REGION Network 23: Buzzer
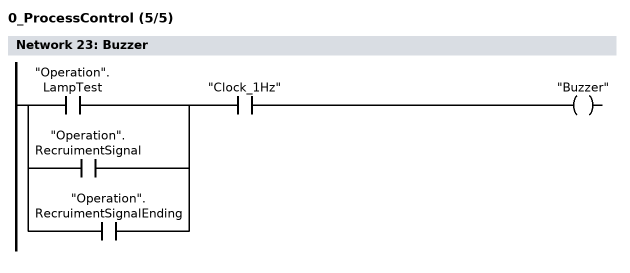
   RUNG wire#powerrail
      Contact( "Operation".LampTest )
      wire#w1
      Contact( "Clock_1Hz" )
      Coil( "Buzzer" )
   END_RUNG
   RUNG wire#powerrail
      Contact( "Operation".RecruimentSignal )
   END_RUNG wire#w1
   RUNG wire#powerrail
      Contact( "Operation".RecruimentSignalEnding )
   END_RUNG wire#w1
   // the same network as SCL:
   "Buzzer" := ("Operation".LampTest OR "Operation".RecruimentSignal OR "Operation".RecruimentSignalEnding) AND "Clock_1Hz";
END_REGION
END_FUNCTION_BLOCK

// folder: 5_Library

FUNCTION_BLOCK "DigAlarm"   // FB2000, SCL
TITLE = Digital Alarm
{ S7_Optimized_Access := 'TRUE' }
AUTHOR : JL_Cristobal_2020
VERSION : 0.1
// Digital Alarm supervisor, trigger memory , ack + reset
   VAR_INPUT
      Pulse : Bool;
      ACK : Bool;
      Reset : Bool;
      Funtion : Bool;
      Input : Bool;
   END_VAR
   VAR_OUTPUT
      DisplayOutput : Bool;
      DisplayOutputNeg : Bool;
      InterlockOutput : Bool;
      InterlockOutputNeg : Bool;
   END_VAR
   VAR
      DisplayAlarmMem : Bool;
      ACKMem : Bool;
      InterlockalarmMem : Bool;
      InterlockMem : Bool;
   END_VAR
BEGIN
   //Alarm process

   //TRUE Mode, Positive Signal
   IF #Funtion = 1 THEN

       IF NOT #Input THEN
           #InterlockMem := false;
           #DisplayAlarmMem := true;
           #InterlockalarmMem := true;
       END_IF;

       IF #Input AND #Reset THEN
           #DisplayAlarmMem := false;
       END_IF;

       IF NOT #Input AND #ACK THEN
           #ACKMem := true;
       END_IF;

       IF #Input AND #Reset THEN
           #InterlockMem := true;
           #ACKMem := false;
           #InterlockalarmMem := false;
       END_IF;

   END_IF;

   //FALSE Mode, Negative Signal
   IF #Funtion = 0 THEN

       IF #Input THEN
           #DisplayAlarmMem := true;
           #InterlockalarmMem := true;
           #InterlockMem := false;
       END_IF;

       IF NOT #Input AND #Reset THEN
           #DisplayAlarmMem := false;
       END_IF;

       IF #Input AND #ACK THEN
           #ACKMem := true;
       END_IF;

       IF NOT #Input AND #Reset THEN
           #ACKMem := false;
           #InterlockalarmMem := false;
           #InterlockMem := true;
       END_IF;

   END_IF;


   #DisplayOutput := #DisplayAlarmMem AND ((#Pulse AND NOT #ACKMem) OR #ACKMem);
   #DisplayOutputNeg := NOT (#DisplayAlarmMem AND ((#Pulse AND NOT #ACKMem) OR #ACKMem));
   #InterlockOutput := #InterlockMem;
   #InterlockOutputNeg := NOT #InterlockMem;
END_FUNCTION_BLOCK

FUNCTION_BLOCK "DigAlarmInterlock"   // FB2001, SCL
TITLE = Digital Alarm With Interlock
{ S7_Optimized_Access := 'TRUE' }
AUTHOR : JL_Cristobal_2020
FAMILY : Alarms
VERSION : 0.1
// Digital Alarm supervisor with interlock signal, trigger memory , ack + reset
   VAR_INPUT
      Pulse : Bool;
      ACK : Bool;
      Reset : Bool;
      Function : Int;
      AlarmInput : Bool;
      SupervisorInput : Bool;
      StartInput : Bool;
      Delay : Time;
   END_VAR
   VAR_OUTPUT
      DisplayOutput : Bool;
      DisplayOutputNeg : Bool;
      InterlockOutput : Bool;
      InterlockOutputNeg : Bool;
      SupervisorOutput : Bool;
      TimeElapsed : Time;
   END_VAR
   VAR RETAIN
      DisplayAlarmMem : Bool;
      ACKMem : Bool;
      InterlockalarmMem : Bool;
      InterlockMem : Bool;
   END_VAR
   VAR
      EndSPVMem : Bool;
   END_VAR
   VAR RETAIN
      SPVMem : Bool;
   END_VAR
BEGIN
   (*GESTION DE LA ALARMA*)

   //TRUE MODE, ACTIVE OK
   IF #Function = 1 OR #Function=3 THEN

       IF NOT #AlarmInput THEN
           #InterlockMem := false;
           #DisplayAlarmMem := true;
           #InterlockalarmMem := true;
       END_IF;

       IF #AlarmInput AND #Reset THEN
           #DisplayAlarmMem := false;
       END_IF;

       IF NOT #AlarmInput AND #ACK THEN
           #ACKMem := true;
       END_IF;

       IF #AlarmInput AND #Reset THEN
           #InterlockMem := true;
           #ACKMem := false;
           #InterlockalarmMem := false;
       END_IF;

   END_IF;

   //FALSE MODE, PASIVE OK
   IF #Function = 0 OR #Function=2 THEN

       IF #AlarmInput THEN
           #DisplayAlarmMem := true;
           #InterlockalarmMem := true;
           #InterlockMem := false;
       END_IF;

       IF NOT #AlarmInput AND #Reset THEN
           #DisplayAlarmMem := false;
       END_IF;

       IF #AlarmInput AND #ACK THEN
           #ACKMem := true;
       END_IF;

       IF NOT #AlarmInput AND #Reset THEN
           #ACKMem := false;
           #InterlockalarmMem := false;
           #InterlockMem := true;
       END_IF;
   END_IF;

   //SUPERVISION CONTROL
   IF #Function = 0 OR #Function = 1 THEN
       IF #StartInput THEN
           "IEC_Timer_0_DB_SPV".TON(IN := #StartInput,
                                    PT := #Delay,
                                    Q => #EndSPVMem,
                                    ET => #TimeElapsed);
           IF #EndSPVMem AND NOT #SupervisorInput THEN
               #SPVMem := 1;
           END_IF;
       ELSE
           #SPVMem := 0;
       END_IF;
   END_IF;


   #DisplayOutput := #DisplayAlarmMem AND ((#Pulse AND NOT #ACKMem) OR #ACKMem);
   #DisplayOutputNeg := NOT (#DisplayAlarmMem AND ((#Pulse AND NOT #ACKMem) OR #ACKMem));
   #InterlockOutput := #InterlockMem;
   #InterlockOutputNeg := NOT #InterlockMem;
END_FUNCTION_BLOCK

FUNCTION_BLOCK "DirectAnalog"   // FB2002, SCL
TITLE = Analog Alarm INT
{ S7_Optimized_Access := 'FALSE' }
AUTHOR : JL_Cristobal_2020
VERSION : 0.1
// Analog (int) Alarm supervisor, trigger memory , ack + reset. Prealarm and alarm for HI and LOW levels
   VAR_INPUT
      Pulse : Bool;
      ACK : Bool;
      Reset : Bool;
      Interlock : Bool;
      Delay : Time;
      Factor : Real;
      AnalogInput : Int;
      SetpointPreAlarmHI : Real;
      SetpointAlarmHI : Real;
      SetpointPreAlarmLOW : Real;
      SetpointAlarmLOW : Real;
      HysteresisHI : Real;
      HysteresisLOW : Real;
   END_VAR
   VAR_OUTPUT
      DisplayPreAlarmHI : Bool;
      InterlockPreAlarmHI : Bool;
      DisplayAlarmHI : Bool;
      InterlockAlarmHI : Bool;
      DisplayPreAlarmLOW : Bool;
      InterlockPreAlarmLOW : Bool;
      DisplayAlarmLOW : Bool;
      InterlockAlarmLOW : Bool;
      CovertedOutput : Real;
      CalcHysterisHI : Real;
      CalcHysteresisLOW : Real;
      DATOS : Struct
         InterlockPreAlarmHI : Bool;
         InterlockAlarmHI : Bool;
         InterlockPreAlarmLOW : Bool;
         InterlockAlarmLOW : Bool;
         CovertedOutput : Real;
         Error : Bool;
      END_STRUCT;
   END_VAR
   VAR
      MemDisplayPreAlarmHI : Bool;
      MemInterlockPreAlarmHI : Bool;
      MemDisplayAlarmHI : Bool;
      MemInterlockAlarmHI : Bool;
      MemDisplayPreAlarmLOW : Bool;
      MemInterlockPreAlarmLOW : Bool;
      MemDisplayAlarmLOW : Bool;
      MemInterlockAlarmLOW : Bool;
   END_VAR
BEGIN
   //Unit conversion
   #CovertedOutput := #AnalogInput/#Factor;

   //Prealarm HI
   //Set PreAlarm
   IF #Interlock AND (#CovertedOutput >= #SetpointPreAlarmHI) THEN
     #InterlockPreAlarmHI := false;
     #MemDisplayPreAlarmHI := true;
   END_IF;
   //ACK
   IF (#MemDisplayPreAlarmHI OR NOT #MemInterlockPreAlarmHI) AND #ACK THEN
     #MemInterlockPreAlarmHI := true;
   END_IF;
   //Reset
   IF(#CovertedOutput < (#SetpointPreAlarmHI - #HysteresisHI)) THEN
     #InterlockPreAlarmHI := true;
     #MemDisplayPreAlarmHI := false;
     #MemInterlockPreAlarmHI := false;
   END_IF;
   //Display Output
   #DisplayPreAlarmHI := NOT #InterlockPreAlarmHI AND ((#Pulse AND NOT #MemInterlockPreAlarmHI) OR #MemInterlockPreAlarmHI);

   //Alarm HI
   //Set Alarm HI
   IF #Interlock AND (#CovertedOutput >= #SetpointAlarmHI) THEN
       #InterlockAlarmHI := false;
     #MemDisplayAlarmHI := true;
   END_IF;
   //ACK
   IF (#MemDisplayAlarmHI OR NOT #MemInterlockAlarmHI) AND #ACK THEN
     #MemInterlockAlarmHI := true;
   END_IF;
   //Reset
   IF(#CovertedOutput < (#SetpointAlarmHI - #HysteresisHI)) THEN
     #InterlockAlarmHI := true;
     #MemDisplayAlarmHI := false;
     #MemInterlockAlarmHI := false;
   END_IF;
   //Display Output
   #DisplayAlarmHI := NOT #InterlockAlarmHI AND ((#Pulse AND NOT #MemInterlockAlarmHI) OR #MemInterlockAlarmHI);
   #CalcHysterisHI := #SetpointAlarmHI - #HysteresisHI;

   //Prealarm LOW
   //Set PreAlarm LOW
   IF #Interlock AND (#CovertedOutput <= #SetpointPreAlarmLOW) THEN
     #InterlockPreAlarmLOW := false;
     #MemDisplayPreAlarmLOW := true;
   END_IF;
   //ACK
   IF (#MemDisplayPreAlarmLOW OR NOT #MemInterlockPreAlarmLOW) AND #ACK THEN
     #MemInterlockPreAlarmLOW := true;
   END_IF;
   //Reset
   IF (#CovertedOutput > (#SetpointPreAlarmLOW + #HysteresisLOW)) THEN
     #InterlockPreAlarmLOW := true;
     #MemDisplayPreAlarmLOW := false;
     #MemInterlockPreAlarmLOW := false;
   END_IF;
   //Display Output
   #DisplayPreAlarmLOW := NOT #InterlockPreAlarmLOW AND ((#Pulse AND NOT #MemInterlockPreAlarmLOW) OR #MemInterlockPreAlarmLOW);

   //Alarm LOW
   //Set Alarm LOW
   IF #Interlock AND (#CovertedOutput <= #SetpointAlarmLOW) THEN
     #InterlockAlarmLOW := false;
     #MemDisplayAlarmLOW := true;
   END_IF;
   //ACK
   IF (#MemDisplayAlarmLOW OR NOT #MemInterlockAlarmLOW )AND #ACK THEN
     #MemInterlockAlarmLOW := true;
   END_IF;
   //Reset
   IF (#CovertedOutput > (#SetpointAlarmLOW + #HysteresisLOW)) THEN
     #InterlockAlarmLOW := true;
     #MemDisplayAlarmLOW := false;
     #MemInterlockAlarmLOW := false;
   END_IF;
   //Display Output
   #DisplayAlarmLOW := NOT #InterlockAlarmLOW AND ((#Pulse AND NOT #MemInterlockAlarmLOW) OR #MemInterlockAlarmLOW);
   #CalcHysteresisLOW := #SetpointAlarmLOW + #HysteresisLOW;

   //Data Output
   #DATOS.InterlockPreAlarmHI := #InterlockPreAlarmHI;
   #DATOS.InterlockAlarmHI := #InterlockAlarmHI;
   #DATOS.InterlockPreAlarmLOW := #InterlockPreAlarmLOW;
   #DATOS.InterlockAlarmLOW := #InterlockAlarmLOW;
   #DATOS.CovertedOutput := #CovertedOutput;
   #DATOS.Error := FALSE;
END_FUNCTION_BLOCK

FUNCTION_BLOCK "DirectAnalogReal"   // FB2003, SCL
TITLE = Analog Alarm REAL
{ S7_Optimized_Access := 'TRUE' }
AUTHOR : JL_Cristobal_2020
VERSION : 0.1
// Analog Alarm (real) supervisor, trigger memory , ack + reset. Prealarm and alarm for HI and LOW levels
   VAR_INPUT
      PULSOS : Bool;
      ENTERADO : Bool;
      REARME : Bool;
      FACTOR : Real;
      ENTRADA_ANALOGICA : Real;
      ValPreALM_SUPERIOR : Real;
      ValALM_SUPERIOR : Real;
      ValPreALM_INFERIOR : Real;
      ValALM_INFERIOR : Real;
      HISTERESIS_SUP : Real;
      HISTERESIS_INF : Real;
   END_VAR
   VAR_OUTPUT
      VIS_PreALM_SUPERIOR : Bool;
      ENC_PreALM_SUPERIOR : Bool;
      VIS_ALM_SUPERIOR : Bool;
      ENC_ALM_SUPERIOR : Bool;
      VIS_PreALM_INFERIOR : Bool;
      ENC_PreALM_INFERIOR : Bool;
      VIS_ALM_INFERIOR : Bool;
      ENC_ALM_INFERIOR : Bool;
      Salida_CONVERTIDA : Real;
      CONS_HIST_SUP : Real;
      CONS_HIST_INF : Real;
      DATOS : Struct
         ENC_PALM_SUP : Bool;
         ENC_ALM_SUP : Bool;
         ENC_PALM_INF : Bool;
         ENC_ALM_INF : Bool;
         VALOR : Real;
         ERROR : Bool;
      END_STRUCT;
   END_VAR
   VAR
      MEM_VIS_PreALM_SUPERIOR : Bool;
      MEM_ENC_PreALM_SUPERIOR : Bool;
      MEM_VIS_ALM_SUPERIOR : Bool;
      MEM_ENC_ALM_SUPERIOR : Bool;
      MEM_VIS_PreALM_INFERIOR : Bool;
      MEM_ENC_PreALM_INFERIOR : Bool;
      MEM_VIS_ALM_INFERIOR : Bool;
      MEM_ENC_ALM_INFERIOR : Bool;
   END_VAR
BEGIN
   (****Conversion de Unidades****)
   #Salida_CONVERTIDA := #ENTRADA_ANALOGICA / #FACTOR;

   (****Prealarma Superior****)
   (*DISPARO DE LA ALARMA*)
   IF (#Salida_CONVERTIDA >= #ValPreALM_SUPERIOR) THEN
       #ENC_PreALM_SUPERIOR := false;
       #MEM_VIS_PreALM_SUPERIOR := true;
   END_IF;
   (*ENTERADO DEFECTO*)
   IF #MEM_VIS_PreALM_SUPERIOR AND #ENTERADO THEN
       #MEM_ENC_PreALM_SUPERIOR := true;
   END_IF;
   (*REARME DEFECTO*)
   IF #REARME AND (#Salida_CONVERTIDA < (#ValPreALM_SUPERIOR - #HISTERESIS_SUP)) THEN
       #ENC_PreALM_SUPERIOR := true;
       #MEM_VIS_PreALM_SUPERIOR := false;
       #MEM_ENC_PreALM_SUPERIOR := false;
   END_IF;
   (*SALIDA VISUALIZACION*)
   #VIS_PreALM_SUPERIOR := NOT #ENC_PreALM_SUPERIOR AND ((#PULSOS AND NOT #MEM_ENC_PreALM_SUPERIOR) OR #MEM_ENC_PreALM_SUPERIOR);

   (****Alarma Superior****)
   (*DISPARO DE LA ALARMA*)
   IF (#Salida_CONVERTIDA >= #ValALM_SUPERIOR) THEN
       #ENC_ALM_SUPERIOR := false;
       #MEM_VIS_ALM_SUPERIOR := true;
   END_IF;
   (*ENTERADO DEFECTO*)
   IF #MEM_VIS_ALM_SUPERIOR AND #ENTERADO THEN
       #MEM_ENC_ALM_SUPERIOR := true;
   END_IF;
   (*REARME DEFECTO*)
   IF #REARME AND (#Salida_CONVERTIDA < (#ValALM_SUPERIOR - #HISTERESIS_SUP)) THEN
       #ENC_ALM_SUPERIOR := true;
       #MEM_VIS_ALM_SUPERIOR := false;
       #MEM_ENC_ALM_SUPERIOR := false;
   END_IF;
   (*SALIDA VISUALIZACION*)
   #VIS_ALM_SUPERIOR := NOT #ENC_ALM_SUPERIOR AND ((#PULSOS AND NOT #MEM_ENC_ALM_SUPERIOR) OR #MEM_ENC_ALM_SUPERIOR);
   #CONS_HIST_SUP := #ValALM_SUPERIOR - #HISTERESIS_SUP;

   (****Prealarma Inferior****)
   (*DISPARO DE LA ALARMA*)
   IF (#Salida_CONVERTIDA <= #ValPreALM_INFERIOR) THEN
       #ENC_PreALM_INFERIOR := false;
       #MEM_VIS_PreALM_INFERIOR := true;
   END_IF;
   (*ENTERADO DEFECTO*)
   IF #MEM_VIS_PreALM_INFERIOR AND #ENTERADO THEN
       #MEM_ENC_PreALM_INFERIOR := true;
   END_IF;
   (*REARME DEFECTO*)
   IF #REARME AND (#Salida_CONVERTIDA > (#ValPreALM_INFERIOR + #HISTERESIS_INF)) THEN
       #ENC_PreALM_INFERIOR := true;
       #MEM_VIS_PreALM_INFERIOR := false;
       #MEM_ENC_PreALM_INFERIOR := false;
   END_IF;
   (*SALIDA VISUALIZACION*)
   #VIS_PreALM_INFERIOR := NOT #ENC_PreALM_INFERIOR AND ((#PULSOS AND NOT #MEM_ENC_PreALM_INFERIOR) OR #MEM_ENC_PreALM_INFERIOR);

   (****Alarma Inferior****)
   (*DISPARO DE LA ALARMA*)
   IF (#Salida_CONVERTIDA <= #ValALM_INFERIOR) THEN
       #ENC_ALM_INFERIOR := false;
       #MEM_VIS_ALM_INFERIOR := true;
   END_IF;
   (*ENTERADO DEFECTO*)
   IF #MEM_VIS_ALM_INFERIOR AND #ENTERADO THEN
       #MEM_ENC_ALM_INFERIOR := true;
   END_IF;
   (*REARME DEFECTO*)
   IF #REARME AND (#Salida_CONVERTIDA > (#ValALM_INFERIOR + #HISTERESIS_INF)) THEN
       #ENC_ALM_INFERIOR := true;
       #MEM_VIS_ALM_INFERIOR := false;
       #MEM_ENC_ALM_INFERIOR := false;
   END_IF;
   (*SALIDA VISUALIZACION*)
   #VIS_ALM_INFERIOR := NOT #ENC_ALM_INFERIOR AND ((#PULSOS AND NOT #MEM_ENC_ALM_INFERIOR) OR #MEM_ENC_ALM_INFERIOR);
   #CONS_HIST_INF := #ValALM_INFERIOR + #HISTERESIS_INF;

   (****SALIDA DATOS****)
   #DATOS.ENC_PALM_SUP := #ENC_PreALM_SUPERIOR;
   #DATOS.ENC_ALM_SUP := #ENC_ALM_SUPERIOR;
   #DATOS.ENC_PALM_INF := #ENC_PreALM_INFERIOR;
   #DATOS.ENC_ALM_INF := #ENC_ALM_INFERIOR;
   #DATOS.VALOR := #Salida_CONVERTIDA;
   #DATOS.ERROR := FALSE;
END_FUNCTION_BLOCK

FUNCTION_BLOCK "Pack_16B"   // FB2004, SCL
TITLE = Pack 16 Digital Alarms in one WORD for HMI transmission
{ S7_Optimized_Access := 'FALSE' }
AUTHOR : JL_Cristobal_2020
VERSION : 0.1
// Pack 16 Digital Alarms in one WORD for HMI transmission, swapping bytes for HMI representation
   VAR_INPUT
      Alarm_0 : Bool;
      Alarm_1 : Bool;
      Alarm_2 : Bool;
      Alarm_3 : Bool;
      Alarm_4 : Bool;
      Alarm_5 : Bool;
      Alarm_6 : Bool;
      Alarm_7 : Bool;
      Alarm_8 : Bool;
      Alarm_9 : Bool;
      Alarm_10 : Bool;
      Alarm_11 : Bool;
      Alarm_12 : Bool;
      Alarm_13 : Bool;
      Alarm_14 : Bool;
      Alarm_15 : Bool;
   END_VAR
   VAR_OUTPUT
      Alarmas_word : Word;
      Alarmas AT Alarmas_word : Array[0..15] of Bool;
   END_VAR
BEGIN
   #Alarmas[0] := NOT #Alarm_8;
   #Alarmas[1] := NOT #Alarm_9;
   #Alarmas[2] := NOT #Alarm_10;
   #Alarmas[3] := NOT #Alarm_11;
   #Alarmas[4] := NOT #Alarm_12;
   #Alarmas[5] := NOT #Alarm_13;
   #Alarmas[6] := NOT #Alarm_14;
   #Alarmas[7] := NOT #Alarm_15;
   #Alarmas[8] := NOT #Alarm_0;
   #Alarmas[9] := NOT #Alarm_1;
   #Alarmas[10] := NOT #Alarm_2;
   #Alarmas[11] := NOT #Alarm_3;
   #Alarmas[12] := NOT #Alarm_4;
   #Alarmas[13] := NOT #Alarm_5;
   #Alarmas[14] := NOT #Alarm_6;
   #Alarmas[15] := NOT #Alarm_7;
END_FUNCTION_BLOCK

FUNCTION_BLOCK "Pack_32B"   // FB2005, SCL
TITLE = Pack 32 Digital Alarms in one DWORD for HMI
{ S7_Optimized_Access := 'TRUE' }
AUTHOR : JL_Cristobal_2020
VERSION : 0.1
// Pack 32 Digital Alarms in one DWORD for HMI transmission, swapping bytes for HMI representation
   VAR_INPUT
      ENTRADA_1 : Bool;
      ENTRADA_2 : Bool;
      ENTRADA_3 : Bool;
      ENTRADA_4 : Bool;
      ENTRADA_5 : Bool;
      ENTRADA_6 : Bool;
      ENTRADA_7 : Bool;
      ENTRADA_8 : Bool;
      ENTRADA_9 : Bool;
      ENTRADA_10 : Bool;
      ENTRADA_11 : Bool;
      ENTRADA_12 : Bool;
      ENTRADA_13 : Bool;
      ENTRADA_14 : Bool;
      ENTRADA_15 : Bool;
      ENTRADA_16 : Bool;
      ENTRADA_17 : Bool;
      ENTRADA_18 : Bool;
      ENTRADA_19 : Bool;
      ENTRADA_20 : Bool;
      ENTRADA_21 : Bool;
      ENTRADA_22 : Bool;
      ENTRADA_23 : Bool;
      ENTRADA_24 : Bool;
      ENTRADA_25 : Bool;
      ENTRADA_26 : Bool;
      ENTRADA_27 : Bool;
      ENTRADA_28 : Bool;
      ENTRADA_29 : Bool;
      ENTRADA_30 : Bool;
      ENTRADA_31 : Bool;
      ENTRADA_32 : Bool;
   END_VAR
   VAR_OUTPUT
      SALIDA : Struct
         SALIDA_1 : Bool;
         SALIDA_2 : Bool;
         SALIDA_3 : Bool;
         SALIDA_4 : Bool;
         SALIDA_5 : Bool;
         SALIDA_6 : Bool;
         SALIDA_7 : Bool;
         SALIDA_8 : Bool;
         SALIDA_9 : Bool;
         SALIDA_10 : Bool;
         SALIDA_11 : Bool;
         SALIDA_12 : Bool;
         SALIDA_13 : Bool;
         SALIDA_14 : Bool;
         SALIDA_15 : Bool;
         SALIDA_16 : Bool;
         SALIDA_17 : Bool;
         SALIDA_18 : Bool;
         SALIDA_19 : Bool;
         SALIDA_20 : Bool;
         SALIDA_21 : Bool;
         SALIDA_22 : Bool;
         SALIDA_23 : Bool;
         SALIDA_24 : Bool;
         SALIDA_25 : Bool;
         SALIDA_26 : Bool;
         SALIDA_27 : Bool;
         SALIDA_28 : Bool;
         SALIDA_29 : Bool;
         SALIDA_30 : Bool;
         SALIDA_31 : Bool;
         SALIDA_32 : Bool;
      END_STRUCT;
   END_VAR
BEGIN
   #SALIDA.SALIDA_1 := #ENTRADA_1;
   #SALIDA.SALIDA_2 := #ENTRADA_2;
   #SALIDA.SALIDA_3 := #ENTRADA_3;
   #SALIDA.SALIDA_4 := #ENTRADA_4;
   #SALIDA.SALIDA_5 := #ENTRADA_5;
   #SALIDA.SALIDA_6 := #ENTRADA_6;
   #SALIDA.SALIDA_7 := #ENTRADA_7;
   #SALIDA.SALIDA_8 := #ENTRADA_8;
   #SALIDA.SALIDA_9 := #ENTRADA_9;
   #SALIDA.SALIDA_10 := #ENTRADA_10;
   #SALIDA.SALIDA_11 := #ENTRADA_11;
   #SALIDA.SALIDA_12 := #ENTRADA_12;
   #SALIDA.SALIDA_13 := #ENTRADA_13;
   #SALIDA.SALIDA_14 := #ENTRADA_14;
   #SALIDA.SALIDA_15 := #ENTRADA_15;
   #SALIDA.SALIDA_16 := #ENTRADA_16;
   #SALIDA.SALIDA_17 := #ENTRADA_17;
   #SALIDA.SALIDA_18 := #ENTRADA_18;
   #SALIDA.SALIDA_19 := #ENTRADA_19;
   #SALIDA.SALIDA_20 := #ENTRADA_20;
   #SALIDA.SALIDA_21 := #ENTRADA_21;
   #SALIDA.SALIDA_22 := #ENTRADA_22;
   #SALIDA.SALIDA_23 := #ENTRADA_23;
   #SALIDA.SALIDA_24 := #ENTRADA_24;
   #SALIDA.SALIDA_25 := #ENTRADA_25;
   #SALIDA.SALIDA_26 := #ENTRADA_26;
   #SALIDA.SALIDA_27 := #ENTRADA_27;
   #SALIDA.SALIDA_28 := #ENTRADA_28;
   #SALIDA.SALIDA_29 := #ENTRADA_29;
   #SALIDA.SALIDA_30 := #ENTRADA_30;
   #SALIDA.SALIDA_31 := #ENTRADA_31;
   #SALIDA.SALIDA_32 := #ENTRADA_32;
END_FUNCTION_BLOCK

FUNCTION_BLOCK "PIDSwitch"   // FB2006, SCL
TITLE = PID Input Parameters Switch
{ S7_Optimized_Access := 'TRUE' }
AUTHOR : JL_Cristobal_2020
VERSION : 0.1
// PID input parameters SWITCH, for multiple secuences
   VAR_INPUT
      A_Setpoint : Real;
      A_Input : Real;
      A_InputPER : Real;
      A_ErrorACK : Bool;
      A_Reset : Bool;
      A_ModeActivate : Bool;
      A_Mode : Int;
      A_Interlock : Bool;
      B_Setpoint : Real;
      B_Input : Real;
      B_InputPER : Real;
      B_ErrorACK : Bool;
      B_Reset : Bool;
      B_ModeActivate : Bool;
      B_Mode : Int;
      B_Interlock : Bool;
      C_Setpoint : Real;
      C_Input : Real;
      C_InputPER : Real;
      C_ErrorACK : Bool;
      C_Reset : Bool;
      C_ModeActivate : Bool;
      C_Mode : Int;
      C_Interlock : Bool;
      D_Setpoint : Real;
      D_Input : Real;
      D_InputPER : Real;
      D_ErrorACK : Bool;
      D_Reset : Bool;
      D_ModeActivate : Bool;
      D_Mode : Int;
      D_Interlock : Bool;
      ChannelSelect : Int;
   END_VAR
   VAR_OUTPUT
      Setpoint : Real;
      Input : Real;
      InputPER : Real;
      ErrorACK : Bool;
      Reset : Bool;
      ModeActivate : Bool;
      Mode : Int;
      Interlock : Bool;
   END_VAR
BEGIN
   CASE #ChannelSelect OF
       1:  // Statement section case 1
           #Setpoint := #A_Setpoint;
           #Input := #A_Input;
           #InputPER := #A_InputPER;
           #ErrorACK := #A_ErrorACK;
           #Reset := #A_Reset;
           #ModeActivate := #A_ModeActivate;
           #Mode := #A_Mode;
       2:  // Statement section case 2
           #Setpoint := #B_Setpoint;
           #Input := #B_Input;
           #InputPER := #B_InputPER;
           #ErrorACK := #B_ErrorACK;
           #Reset := #B_Reset;
           #ModeActivate := #B_ModeActivate;
           #Mode := #B_Mode;
       3:  // Statement section case 3
           #Setpoint := #C_Setpoint;
           #Input := #C_Input;
           #InputPER := #C_InputPER;
           #ErrorACK := #A_ErrorACK;
           #Reset := #C_Reset;
           #ModeActivate := #C_ModeActivate;
           #Mode := #C_Mode;
       4:  // Statement section case 4
           #Setpoint := #D_Setpoint;
           #Input := #D_Input;
           #InputPER := #D_InputPER;
           #ErrorACK := #D_ErrorACK;
           #Reset := #D_Reset;
           #ModeActivate := #D_ModeActivate;
           #Mode := #D_Mode;
       ELSE  // Statement section ELSE
           #Setpoint := 0.0;
           #Input := 0.0;
           #InputPER := 0.0;
           #ErrorACK := FALSE;
           #Reset := TRUE;
           #ModeActivate := FALSE;
           #Mode := 0;
   END_CASE;
END_FUNCTION_BLOCK

FUNCTION_BLOCK "RatioCalculator"   // FB2007, SCL
TITLE = Ratio Calculator
{ S7_Optimized_Access := 'TRUE' }
AUTHOR : JL_Cristobal_2020
VERSION : 0.1
// Ratio Calculator for relation between Inspiration, Delay and Espiration
   VAR_INPUT
      BPM : Real;
   END_VAR
   VAR_OUTPUT
      CalculatedRatio : Real;
      InspirationTime : Time;
      RestTime : Time;
      EspirationTime : Time;
      DelayTime : Time;
      TotalTime : Time;
   END_VAR
   VAR_IN_OUT
      Inspiration : Real;
      Espiration : Real;
      Delay : Real;
      Rest : Real;
   END_VAR
   VAR
      BPMTimeReal : Real;
      InspTimeReal : Real;
      EspTimeReal : Real;
      DelayTimeReal : Real;
      RestTimeReal : Real;
      TotalTimeReal : Real;
      BPMTimeInt : Int;
      InspTimeInt : Int;
      EspTimeInt : Int;
      DelayTimeInt : Int;
      RestTimeInt : Int;
      TotalTimeInt : Int;
   END_VAR
BEGIN
   //BPM calculator
   #BPMTimeReal:=60.0/#BPM;
   #TotalTimeInt := #BPMTimeReal * 1000;
   #TotalTime := INT_TO_TIME(#TotalTimeInt);

   //Inspiration calculator
   #InspTimeReal := #BPMTimeReal * (#Inspiration/100.0);
   #InspTimeInt := #InspTimeReal * 1000;
   #InspirationTime := INT_TO_TIME(#InspTimeInt);
   IF #Inspiration > 50 THEN
       #Inspiration := 50;
   END_IF;

   //Rest Time
   #Rest := 100.0 - #Inspiration;
   #RestTimeReal := #BPMTimeReal - #InspTimeReal;
   #RestTimeInt := #RestTimeReal * 1000;
   #RestTime := INT_TO_TIME(#RestTimeInt);

   //Espiration Time
   #EspTimeReal:=#BPMTimeReal *(#Espiration/100.0);
   #EspTimeInt := #EspTimeReal * 1000;
   #EspirationTime := INT_TO_TIME(#EspTimeInt);
   IF #Espiration >=50 THEN
       IF #Inspiration >= 50 THEN
           #Espiration := 40;
       ELSE
           #Espiration := 50;
       END_IF;
   END_IF;

   //Delay Time
   #Delay := #Rest - #Espiration;
   #DelayTimeReal := #RestTimeReal - #EspTimeReal;
   #DelayTimeInt := #DelayTimeReal * 1000;
   #DelayTime := INT_TO_TIME(#DelayTimeInt);

   //Total Time
   #TotalTimeReal := #InspTimeReal + #EspTimeReal + #DelayTimeReal;
END_FUNCTION_BLOCK

FUNCTION_BLOCK "VariableSupervisor"   // FB2008, SCL
TITLE = Variable Supervisor
{ S7_Optimized_Access := 'TRUE' }
AUTHOR : JL_Cristobal_2020
VERSION : 0.1
// Dinamic control for settings between limits
   VAR_INPUT
      SetpointIncrement : Bool;
      SetpointDecrement : Bool;
      Max : Real;
      Min : Real;
   END_VAR
   VAR_IN_OUT
      SetpointMax : Real;
      SetpointMin : Real;
      InOutSetpoint : Real;
      InOutAlarmHI : Real;
      InOutPreAlarmHI : Real;
      InOutAlarmLOW : Real;
      InOutPreAlarmLOW : Real;
   END_VAR
   VAR
      SetpointREPlus : Bool;
      SetpointREMinus : Bool;
      SetpointMemPlus : Bool;
      SetpointMemMinus : Bool;
   END_VAR
BEGIN
   //Variable Supervisor

   //Setpoint Increment
   "R_TRIG_DB_Plus"(CLK:=#SetpointIncrement,
                    Q=>#SetpointREPlus);
   IF #SetpointREPlus AND "Clock_1Hz" AND NOT #SetpointMemPlus THEN
       #InOutSetpoint := #InOutSetpoint + 1;
       #SetpointMemPlus := 1;
   END_IF;
   IF NOT "Clock_1Hz" THEN
       #SetpointMemPlus := 0;
   END_IF;
   IF #InOutSetpoint > #SetpointMax THEN
       #InOutSetpoint := #SetpointMax;
   END_IF;


   //Setpoint Decrement
   "R_TRIG_DB_Minus"(CLK := #SetpointDecrement,
                     Q => #SetpointREMinus);
   IF #SetpointREMinus AND "Clock_1Hz" AND NOT #SetpointMemMinus THEN
       #InOutSetpoint := #InOutSetpoint - 1;
       #SetpointMemMinus := 1;
   END_IF;
   IF NOT "Clock_1Hz" THEN
       #SetpointMemMinus := 0;
   END_IF;
   IF #InOutSetpoint < #SetpointMin THEN
       #InOutSetpoint := #SetpointMin;
   END_IF;

   //MAX Control
   IF #InOutSetpoint > #SetpointMax THEN
       #InOutSetpoint := #SetpointMax;
   END_IF;
   IF #SetpointMax > #Max THEN
       #SetpointMax := #Max;
   END_IF;
   IF #SetpointMax < #SetpointMin THEN
       #SetpointMax := #SetpointMin+1;
   END_IF;

   //MAX Alarm Control
   IF #InOutAlarmHI > #SetpointMax THEN
       #InOutAlarmHI := #SetpointMax;
   END_IF;
   IF #InOutAlarmHI < #SetpointMin THEN
       #InOutAlarmHI := #SetpointMin +2;
   END_IF;
   //MAX PreAlarm Control
   IF #InOutPreAlarmHI > #SetpointMax OR #InOutPreAlarmHI >=#InOutAlarmHI OR #InOutPreAlarmHI < #SetpointMin THEN
       #InOutPreAlarmHI := #InOutAlarmHI-1;
   END_IF;

   //MIN Control
   IF #InOutSetpoint < #SetpointMin THEN
       #InOutSetpoint := #SetpointMin;
   END_IF;
   IF #SetpointMin < #Min THEN
       #SetpointMin := #Min;
   END_IF;
   IF #SetpointMin >#SetpointMax THEN
       #SetpointMin := #SetpointMax -1 ;
   END_IF;

   //MIN Alarm Control
   IF #InOutAlarmLOW < #SetpointMin THEN
       #InOutAlarmLOW := #SetpointMin;
   END_IF;
   IF #InOutAlarmLOW > #SetpointMax THEN
       #InOutAlarmLOW := #SetpointMax - 2;
   END_IF;

   //MIN PreAlarm Control
   IF #InOutPreAlarmLOW < #SetpointMin OR #InOutAlarmLOW <=  #InOutAlarmLOW  OR #InOutPreAlarmLOW > #SetpointMax THEN
       #InOutPreAlarmLOW := #InOutAlarmLOW+1;
   END_IF;
END_FUNCTION_BLOCK

(* ===== HMI "HMI_RT_1" =====
system functions are stored by id; their names below are inferred from use
connection "HMI_Conexión_1": ETHERNET, S7_1200_OMS

HMI tags "Tabla de variables estándar"
   "OperatingParameters_TidalVolumenMax" : Real = PLC OperatingParameters.TidalVolumenMax, 100 ms
   "OperatingParameters_TidalVolumenSetpoint" : Real = PLC OperatingParameters.TidalVolumenSetpoint, 100 ms
   "OperatingParameters_TidalVolumenMin" : Real = PLC OperatingParameters.TidalVolumenMin, 100 ms
   "OperatingParameters_PlateauMax" : Real = PLC OperatingParameters.PlateauMax, 100 ms
   "OperatingParameters_PlateauSetpoint" : Real = PLC OperatingParameters.PlateauSetpoint, 100 ms
   "OperatingParameters_PlateauMin" : Real = PLC OperatingParameters.PlateauMin, 100 ms
   "OperatingParameters_PeepMax" : Real = PLC OperatingParameters.PeepMax, 100 ms
   "OperatingParameters_PeepSetpoint" : Real = PLC OperatingParameters.PeepSetpoint, 100 ms
   "OperatingParameters_PeepMin" : Real = PLC OperatingParameters.PeepMin, 100 ms
   "OperatingParameters_FrequencyMax" : Real = PLC OperatingParameters.FrequencyMax, 100 ms
   "OperatingParameters_FrequencySetpoint" : Real = PLC OperatingParameters.FrequencySetpoint, 100 ms
   "OperatingParameters_FrequencyMin" : Real = PLC OperatingParameters.FrequencyMin, 100 ms
   "OperatingParameters_BatteryLevelTrigger" : Real = PLC OperatingParameters.BatteryLevelTrigger, 100 ms
   "Clock_2.5Hz" : Bool = PLC "Clock_2.5Hz" AT %M0.2, 100 ms
   "Clock_1Hz" : Bool = PLC Clock_1Hz AT %M0.5, 100 ms
   "Clock_Byte" : Byte = PLC Clock_Byte AT %MB0, 100 ms
   "System_Byte" : Byte = PLC System_Byte AT %MB1, 100 ms
   "Variable_HMI_1" : Int, internal
   "ServoAlarm" : Bool = PLC ServoAlarm AT %I1.1, 100 ms
   "AlwaysTRUE" : Bool = PLC AlwaysTRUE AT %M1.2, 100 ms
   "OperatingParameters_PipSetpoint" : Real = PLC OperatingParameters.PipSetpoint, 100 ms
   "OperatingParameters_PipMax" : Real = PLC OperatingParameters.PipMax, 100 ms
   "DataValues_PipValue" : Real = PLC DataValues.PipValue, 100 ms
   "OperatingParameters_PipMin" : Real = PLC OperatingParameters.PipMin, 100 ms
   "DataValues_PlateauValue" : Real = PLC DataValues.PlateauValue, 100 ms
   "DataValues_PeepValue" : Real = PLC DataValues.PeepValue, 100 ms
   "DataValues_FrequencyValue" : Real = PLC DataValues.FrequencyValue, 100 ms
   "DataValues_TidalVolumeValue" : Real = PLC DataValues.TidalVolumeValue, 100 ms
   "DataValues_MinumValue" : Real = PLC DataValues.VolumeMinuteValue, 100 ms
   "OperatingParameters_MinimumVolumeMin" : Real = PLC OperatingParameters.VolumeMinMin, 100 ms
   "OperatingParameters_TriggerSetpoint" : Real = PLC OperatingParameters.TriggerSetpoint, 100 ms
   "DataValues_BatteryVoltage" : Real = PLC DataValues.BatteryVoltage, 100 ms
   "DataValues_BatteryCapacity" : Real = PLC DataValues.BatteryCapacity, 100 ms
   "OperatingParameters_MinimumVolumeMax" : Real = PLC OperatingParameters.VolumeMinMax, 100 ms
   "2_PWMValve_Enable" : Bool = PLC "2_PWMValve".Enable, 100 ms
   "2_PWMValve_Frecuency" : DInt = PLC "2_PWMValve".Frecuency, 100 ms
   "2_PWMValve_Duty_Cycle" : Int = PLC "2_PWMValve".Duty_Cycle, 100 ms
   "PatientData_TidalVolume" : Real = PLC PatientData.TidalVolume, 100 ms
   "PatientData_PatientType" : Int = PLC PatientData.PatientType, 100 ms
   "PatientData_PatientHeight" : Real = PLC PatientData.PatientHeight, 100 ms
   "OperatingParameters_PeakPBMinus" : Bool = PLC OperatingParameters.PeakPBMinus, 100 ms
   "OperatingParameters_PeakPBPlus" : Bool = PLC OperatingParameters.PeakPBPlus, 100 ms
   "OperatingParameters_PeepPBMinus" : Bool = PLC OperatingParameters.PeepPBMinus, 100 ms
   "OperatingParameters_PeepPBPlus" : Bool = PLC OperatingParameters.PeepPBPlus, 100 ms
   "OperatingParameters_FrPBMinus" : Bool = PLC OperatingParameters.FrPBMinus, 100 ms
   "OperatingParameters_FrPBPlus" : Bool = PLC OperatingParameters.FrPBPlus, 100 ms
   "OperatingParameters_RecruitmentOn" : Bool = PLC OperatingParameters.RecruitmentOn, 100 ms
   "OperatingParameters_RecruitmentOff" : Bool = PLC OperatingParameters.RecruitmentOff, 100 ms
   "OperatingParameters_RecruitmentElap" : Time = PLC OperatingParameters.RecruitmentElap, 100 ms
   "DateTime_SystemDateRetVal" : Int = PLC DateTime.SystemDateRetVal AT %DB102.DBW0, 100 ms
   "DateTime_SystemDateOut" : DTL = PLC DateTime.SystemDateOut AT %DB102.DBX2.0, 100 ms
   "MotorControl_POWER_Enable" : Bool = PLC MotorControl.POWER_Enable, 100 ms
   "MotorControl_RESET_Execute" : Bool = PLC MotorControl.RESET_Execute, 100 ms
   "MotorControl_HOME_Execute" : Bool = PLC MotorControl.HOME_Execute, 100 ms
   "MotorControl_HOME_Position" : Real = PLC MotorControl.HOME_Position, 100 ms
   "MotorControl_HALT_Execute" : Bool = PLC MotorControl.HALT_Execute, 100 ms
   "MotorControl_Velocity_Execute" : Bool = PLC MotorControl.Velocity_Execute, 100 ms
   "MotorControl_POWER_Error" : Bool = PLC MotorControl.POWER_Error, 100 ms
   "MotorControl_POWER_Status" : Bool = PLC MotorControl.POWER_Status, 100 ms
   "MotorControl_RESET_Done" : Bool = PLC MotorControl.RESET_Done, 100 ms
   "MotorControl_RESET_Error" : Bool = PLC MotorControl.RESET_Error, 100 ms
   "MotorControl_HALT_Done" : Bool = PLC MotorControl.HALT_Done, 100 ms
   "MotorControl_HALT_Error" : Bool = PLC MotorControl.HALT_Error, 100 ms
   "MotorControl_HOME_Done" : Bool = PLC MotorControl.HOME_Done, 100 ms
   "MotorControl_HOME_Error" : Bool = PLC MotorControl.HOME_Error, 100 ms
   "MotorControl_Velocity_invelocity" : Bool = PLC MotorControl.Velocity_invelocity, 100 ms
   "MotorControl_Velocity_Error" : Bool = PLC MotorControl.Velocity_Error, 100 ms
   "MotorControl_Velocity_Velocity" : Real = PLC MotorControl.Velocity_Velocity, 100 ms
   "MotorControl_JOG_Invelocity" : Bool = PLC MotorControl.JOG_Invelocity, 100 ms
   "MotorControl_JOG_Backward" : Bool = PLC MotorControl.JOG_Backward, 100 ms
   "MotorControl_JOG_Error" : Bool = PLC MotorControl.JOG_Error, 100 ms
   "MotorControl_JOG_Forward" : Bool = PLC MotorControl.JOG_Forward, 100 ms
   "MotorControl_Velocity_Current" : Bool = PLC MotorControl.Velocity_Current, 100 ms
   "MotorControl_JOG_Velocity" : Real = PLC MotorControl.JOG_Velocity, 100 ms
   "MotorControl_ABSOLUTE_Position" : Real = PLC MotorControl.ABSOLUTE_Position, 100 ms
   "MotorControl_ABSOLUTE_Velocity" : Real = PLC MotorControl.ABSOLUTE_Velocity, 100 ms
   "MotorControl_RELATIVE_Velocity" : Real = PLC MotorControl.RELATIVE_Velocity, 100 ms
   "MotorControl_RELATIVE_Distance" : Real = PLC MotorControl.RELATIVE_Distance, 100 ms
   "MotorControl_ABSOLUTE_Execute" : Bool = PLC MotorControl.ABSOLUTE_Execute, 100 ms
   "MotorControl_ABSOLUTE_Done" : Bool = PLC MotorControl.ABSOLUTE_Done, 100 ms
   "MotorControl_ABSOLUTE_Error" : Bool = PLC MotorControl.ABSOLUTE_Error, 100 ms
   "MotorControl_RELATIVE_Done" : Bool = PLC MotorControl.RELATIVE_Done, 100 ms
   "MotorControl_RELATIVE_Error" : Bool = PLC MotorControl.RELATIVE_Error, 100 ms
   "MotorControl_RELATIVE_Execute" : Bool = PLC MotorControl.RELATIVE_Execute, 100 ms
   "2_PWMValve_Status" : Int = PLC "2_PWMValve".Status, 100 ms
   "2_PWMValve_Busy" : Bool = PLC "2_PWMValve".Busy, 100 ms
   "Alarm0Pack16B_Alarmas_word" : Word = PLC Alarm0Pack16B.Alarmas_word AT %DB300.DBW2, 100 ms
   "Alarm1Pack16B_Alarmas_word" : Word = PLC Alarm1Pack16B.Alarmas_word AT %DB301.DBW2, 100 ms
   "Alarm2Pack16B_Alarmas_word" : Word = PLC Alarm2Pack16B.Alarmas_word AT %DB302.DBW2, 100 ms
   "Alarm3Pack16B_Alarmas_word" : Word = PLC Alarm3Pack16B.Alarmas_word AT %DB303.DBW2, 100 ms
   "OperatingParameters_RecruitmentRunning" : Bool = PLC OperatingParameters.RecruitmentRunning, 100 ms
   "OperatingParameters_RecruitmentEnding" : Bool = PLC OperatingParameters.RecruitmentEnding, 100 ms
   "PatientData_PatientWeight" : Real = PLC PatientData.PatientWeight, 100 ms
   "PatientData_TimeStart" : Time_Of_Day = PLC PatientData.TimeStart, 100 ms
   "PatientData_TimeEnd" : Time_Of_Day = PLC PatientData.TimeEnd, 100 ms
   "OperatingParameters_MinimumVolumeSetpoint" : Real = PLC OperatingParameters.VolumeMinSetpoint, 100 ms
   "DataValues_Trigger" : Real = PLC DataValues.Trigger, 100 ms
   "OperatingParameters_Trigger" : Bool = PLC OperatingParameters.Trigger, 100 ms
   "OperatingParameters_RecruitmentMem" : Bool = PLC OperatingParameters.RecruitmentMem, 100 ms
   "OperatingParameters_RecruitmentEnd" : Bool = PLC OperatingParameters.RecruitmentEnd, 100 ms
   "DateTime_LocalDateOut" : DTL = PLC DateTime.LocalDateOut AT %DB102.DBX16.0, 100 ms
   "PIDData_ChannelSelect" : Int = PLC PIDData.ChannelSelect, 100 ms
   "Alarm1Pack16B_Alarm_1" : Bool = PLC Alarm1Pack16B.Alarm_1 AT %DB301.DBX0.1, 100 ms
   "Alarm1Pack16B_Alarm_5" : Bool = PLC Alarm1Pack16B.Alarm_5 AT %DB301.DBX0.5, 100 ms
   "Alarm1Pack16B_Alarm_9" : Bool = PLC Alarm1Pack16B.Alarm_9 AT %DB301.DBX1.1, 100 ms
   "Alarm1Pack16B_Alarm_13" : Bool = PLC Alarm1Pack16B.Alarm_13 AT %DB301.DBX1.5, 100 ms
   "Alarm2Pack16B_Alarm_1" : Bool = PLC Alarm2Pack16B.Alarm_1 AT %DB302.DBX0.1, 100 ms
   "Alarm2Pack16B_Alarm_5" : Bool = PLC Alarm2Pack16B.Alarm_5 AT %DB302.DBX0.5, 100 ms
   "Alarm1Pack16B_Alarm_3" : Bool = PLC Alarm1Pack16B.Alarm_3 AT %DB301.DBX0.3, 100 ms
   "Alarm1Pack16B_Alarm_7" : Bool = PLC Alarm1Pack16B.Alarm_7 AT %DB301.DBX0.7, 100 ms
   "Alarm1Pack16B_Alarm_11" : Bool = PLC Alarm1Pack16B.Alarm_11 AT %DB301.DBX1.3, 100 ms
   "Alarm1Pack16B_Alarm_15" : Bool = PLC Alarm1Pack16B.Alarm_15 AT %DB301.DBX1.7, 100 ms
   "Alarm2Pack16B_Alarm_3" : Bool = PLC Alarm2Pack16B.Alarm_3 AT %DB302.DBX0.3, 100 ms
   "Alarm2Pack16B_Alarm_7" : Bool = PLC Alarm2Pack16B.Alarm_7 AT %DB302.DBX0.7, 100 ms
   "Alarm1Pack16B_Alarm_0" : Bool = PLC Alarm1Pack16B.Alarm_0 AT %DB301.DBX0.0, 100 ms
   "Alarm1Pack16B_Alarm_2" : Bool = PLC Alarm1Pack16B.Alarm_2 AT %DB301.DBX0.2, 100 ms
   "Alarm1Pack16B_Alarm_4" : Bool = PLC Alarm1Pack16B.Alarm_4 AT %DB301.DBX0.4, 100 ms
   "Alarm1Pack16B_Alarm_6" : Bool = PLC Alarm1Pack16B.Alarm_6 AT %DB301.DBX0.6, 100 ms
   "Alarm1Pack16B_Alarm_8" : Bool = PLC Alarm1Pack16B.Alarm_8 AT %DB301.DBX1.0, 100 ms
   "Alarm1Pack16B_Alarm_10" : Bool = PLC Alarm1Pack16B.Alarm_10 AT %DB301.DBX1.2, 100 ms
   "Alarm1Pack16B_Alarm_12" : Bool = PLC Alarm1Pack16B.Alarm_12 AT %DB301.DBX1.4, 100 ms
   "Alarm1Pack16B_Alarm_14" : Bool = PLC Alarm1Pack16B.Alarm_14 AT %DB301.DBX1.6, 100 ms
   "Alarm2Pack16B_Alarm_0" : Bool = PLC Alarm2Pack16B.Alarm_0 AT %DB302.DBX0.0, 100 ms
   "Alarm2Pack16B_Alarm_2" : Bool = PLC Alarm2Pack16B.Alarm_2 AT %DB302.DBX0.2, 100 ms
   "Alarm2Pack16B_Alarm_4" : Bool = PLC Alarm2Pack16B.Alarm_4 AT %DB302.DBX0.4, 100 ms
   "Alarm2Pack16B_Alarm_6" : Bool = PLC Alarm2Pack16B.Alarm_6 AT %DB302.DBX0.6, 100 ms
   "ProcessData_PpipSetpointAlarmHI" : Real = PLC ProcessData.PpipSetpointAlarmHI, 100 ms
   "ProcessData_PipSetpointPreAlarmHI" : Real = PLC ProcessData.PipSetpointPreAlarmHI, 100 ms
   "ProcessData_PipSetpointAlarmLOW" : Real = PLC ProcessData.PipSetpointAlarmLOW, 100 ms
   "ProcessData_PipSetpointPreAlarmLOW" : Real = PLC ProcessData.PipSetpointPreAlarmLOW, 100 ms
   "ProcessData_PlateauSetpointAlarmHI" : Real = PLC ProcessData.PlateauSetpointAlarmHI, 100 ms
   "ProcessData_PlateauSetpointPreAlarmHI" : Real = PLC ProcessData.PlateauSetpointPreAlarmHI, 100 ms
   "ProcessData_PlateaukSetpointAlarmLOW" : Real = PLC ProcessData.PlateauSetpointAlarmLOW, 100 ms
   "ProcessData_PlateauSetpointPreAlarmLOW" : Real = PLC ProcessData.PlateauSetpointPreAlarmLOW, 100 ms
   "ProcessData_PeepSetpointAlarmHI" : Real = PLC ProcessData.PeepSetpointAlarmHI, 100 ms
   "ProcessData_PeepSetpointPreAlarmHI" : Real = PLC ProcessData.PeepSetpointPreAlarmHI, 100 ms
   "ProcessData_PeepSetpointAlarmLOW" : Real = PLC ProcessData.PeepSetpointAlarmLOW, 100 ms
   "ProcessData_PeepSetpointPreAlarmLOW" : Real = PLC ProcessData.PeepSetpointPreAlarmLOW, 100 ms
   "ProcessData_FrequencySetpointAlarmHI" : Real = PLC ProcessData.FrequencySetpointAlarmHI, 100 ms
   "ProcessData_FrequencySetpointPreAlarmHI" : Real = PLC ProcessData.FrequencySetpointPreAlarmHI, 100 ms
   "ProcessData_FrequencySetpointAlarmLOW" : Real = PLC ProcessData.FrequencySetpointAlarmLOW, 100 ms
   "ProcessData_FrequencySetpointPreAlarmLOW" : Real = PLC ProcessData.FrequencySetpointPreAlarmLOW, 100 ms
   "ProcessData_TidalVolumeSetpointAlarmHI" : Real = PLC ProcessData.TidalVolumeSetpointAlarmHI, 100 ms
   "ProcessData_TidalVolumeSetpointPreAlarmHI" : Real = PLC ProcessData.TidalVolumeSetpointPreAlarmHI, 100 ms
   "ProcessData_TidalVolumeSetpointAlarmLOW" : Real = PLC ProcessData.TidalVolumeSetpointAlarmLOW, 100 ms
   "ProcessData_TidalVolumeSetpointPreAlarmLOW" : Real = PLC ProcessData.TidalVolumeSetpointPreAlarmLOW, 100 ms
   "OperatingParameters_TriggerMax" : Real = PLC OperatingParameters.TriggerMax, 100 ms
   "OperatingParameters_TriggerMin" : Real = PLC OperatingParameters.TriggerMin, 100 ms
   "ProcessData_TriggerVolumeSetpointAlarmHI" : Real = PLC ProcessData.TriggerVolumeSetpointAlarmHI, 100 ms
   "ProcessData_TriggeVolumeSetpointPreAlarmHI" : Real = PLC ProcessData.TriggeVolumeSetpointPreAlarmHI, 100 ms
   "ProcessData_TriggerVolumeSetpointAlarmLOW" : Real = PLC ProcessData.TriggerVolumeSetpointAlarmLOW, 100 ms
   "ProcessData_TriggerVolumeSetpointPreAlarmLOW" : Real = PLC ProcessData.TriggerVolumeSetpointPreAlarmLOW, 100 ms
   "DataValues_AirPressure" : Real = PLC DataValues.AirPressure, 100 ms
   "DataValues_O2Pressure" : Real = PLC DataValues.O2Pressure, 100 ms
   "OperatingParameters_AirSetpoint" : Real = PLC OperatingParameters.AirSetpoint, 100 ms
   "OperatingParameters_O2Setpoint" : Real = PLC OperatingParameters.O2Setpoint, 100 ms
   "OperatingParameters_Air" : Bool = PLC OperatingParameters.Air, 100 ms
   "OperatingParameters_O2" : Bool = PLC OperatingParameters.O2, 100 ms
   "OperatingParameters_HumidifiertElap" : Time = PLC OperatingParameters.HumidifiertElap, 100 ms
   "OperatingParameters_HumidifierTimer" : Time = PLC OperatingParameters.HumidifierTimer, 100 ms
   "OperatingParameters_HumidifiertDuration" : Time = PLC OperatingParameters.HumidifiertDuration, 100 ms
   "DataValues_DrivingPressure" : Real = PLC DataValues.DrivingPressure, 100 ms
   "OperatingParameters_InpirationRatio" : Real = PLC OperatingParameters.InpirationRatio, 100 ms
   "OperatingParameters_EspirationRatio" : Real = PLC OperatingParameters.EspirationRatio, 100 ms
   "OperatingParameters_DelayRatio" : Real = PLC OperatingParameters.DelayRatio, 100 ms
   "OperatingParameters_CalculatedRatio" : Real = PLC OperatingParameters.CalculatedRatio, 100 ms
   "DataValues_TotalTime" : Time = PLC DataValues.TotalTime, 100 ms
   "DataValues_InspirationTime" : Time = PLC DataValues.InspirationTime, 100 ms
   "DataValues_RestTime" : Time = PLC DataValues.RestTime, 100 ms
   "DataValues_EspirationTime" : Time = PLC DataValues.EspirationTime, 100 ms
   "DataValues_DelayTime" : Time = PLC DataValues.DelayTime, 100 ms
   "OperatingParameters_RestRatio" : Real = PLC OperatingParameters.RestRatio, 100 ms
   "TurnAxis_Position" : Real = PLC TurnAxis.Position, 100 ms
   "OperatingParameters_ControlMode" : Int = PLC OperatingParameters.ControlMode, 100 ms
   "AlarmsRaw_PipDisplayAlarmHI" : Bool = PLC AlarmsRaw.PipDisplayAlarmHI, 100 ms
   "AlarmsRaw_PipDisplayPreAlarmHI" : Bool = PLC AlarmsRaw.PipDisplayPreAlarmHI, 100 ms
   "AlarmsRaw_PipDisplayPreAlarmLOW" : Bool = PLC AlarmsRaw.PipDisplayPreAlarmLOW, 100 ms
   "AlarmsRaw_PipDisplayAlarmLOW" : Bool = PLC AlarmsRaw.PipDisplayAlarmLOW, 100 ms
   "AlarmsRaw_PlateauDisplayAlarmHI" : Bool = PLC AlarmsRaw.PlateauDisplayAlarmHI, 100 ms
   "AlarmsRaw_PlateauDisplayPreAlarmHI" : Bool = PLC AlarmsRaw.PlateauDisplayPreAlarmHI, 100 ms
   "AlarmsRaw_PlateauDisplayPreAlarmLOW" : Bool = PLC AlarmsRaw.PlateauDisplayPreAlarmLOW, 100 ms
   "AlarmsRaw_PlateauDisplayAlarmLOW" : Bool = PLC AlarmsRaw.PlateauDisplayAlarmLOW, 100 ms
   "AlarmsRaw_PeepDisplayAlarmHI" : Bool = PLC AlarmsRaw.PeepDisplayAlarmHI, 100 ms
   "AlarmsRaw_PeepDisplayPreAlarmHI" : Bool = PLC AlarmsRaw.PeepDisplayPreAlarmHI, 100 ms
   "AlarmsRaw_PeepDisplayPreAlarmLOW" : Bool = PLC AlarmsRaw.PeepDisplayPreAlarmLOW, 100 ms
   "AlarmsRaw_PeepDisplayAlarmLOW" : Bool = PLC AlarmsRaw.PeepDisplayAlarmLOW, 100 ms
   "AlarmsRaw_FrequencyDisplayAlarmHI" : Bool = PLC AlarmsRaw.FrequencyDisplayAlarmHI, 100 ms
   "AlarmsRaw_FrequencyDisplayPreAlarmHI" : Bool = PLC AlarmsRaw.FrequencyDisplayPreAlarmHI, 100 ms
   "AlarmsRaw_FrequencyDisplayPreAlarmLOW" : Bool = PLC AlarmsRaw.FrequencyDisplayPreAlarmLOW, 100 ms
   "AlarmsRaw_FrequencyDisplayAlarmLOW" : Bool = PLC AlarmsRaw.FrequencyDisplayAlarmLOW, 100 ms
   "AlarmsRaw_TidalVolumeDisplayAlarmHI" : Bool = PLC AlarmsRaw.TidalVolumeDisplayAlarmHI, 100 ms
   "AlarmsRaw_TidalVolumeDisplayPreAlarmHI" : Bool = PLC AlarmsRaw.TidalVolumeDisplayPreAlarmHI, 100 ms
   "AlarmsRaw_TidalVolumeDisplayPreAlarmLOW" : Bool = PLC AlarmsRaw.TidalVolumeDisplayPreAlarmLOW, 100 ms
   "AlarmsRaw_TidalVolumeDisplayAlarmLOW" : Bool = PLC AlarmsRaw.TidalVolumeDisplayAlarmLOW, 100 ms
   "AlarmsRaw_VolumeMinuteDisplayAlarmHI" : Bool = PLC AlarmsRaw.VolumeMinuteDisplayAlarmHI, 100 ms
   "AlarmsRaw_VolumeMinuteDisplayPreAlarmHI" : Bool = PLC AlarmsRaw.VolumeMinuteDisplayPreAlarmHI, 100 ms
   "AlarmsRaw_VolumeMinuteDisplayPreAlarmLOW" : Bool = PLC AlarmsRaw.VolumeMinuteDisplayPreAlarmLOW, 100 ms
   "AlarmsRaw_VolumeMinuteDisplayAlarmLOW" : Bool = PLC AlarmsRaw.VolumeMinuteDisplayAlarmLOW, 100 ms
   "ProcessData_VolumeMinSetpointAlarmHI" : Real = PLC ProcessData.VolumeMinSetpointAlarmHI, 100 ms
   "ProcessData_VolumeMinSetpointPreAlarmHI" : Real = PLC ProcessData.VolumeMinSetpointPreAlarmHI, 100 ms
   "ProcessData_VolumeMinSetpointPreAlarmLOW" : Real = PLC ProcessData.VolumeMinSetpointPreAlarmLOW, 100 ms
   "ProcessData_VolumeMinSetpointAlarmLOW" : Real = PLC ProcessData.VolumeMinSetpointAlarmLOW, 100 ms
   "AlarmsRaw_TriggerDisplayAlarmHI" : Bool = PLC AlarmsRaw.TriggerDisplayAlarmHI, 100 ms
   "AlarmsRaw_TriggerDisplayPreAlarmHI" : Bool = PLC AlarmsRaw.TriggerDisplayPreAlarmHI, 100 ms
   "AlarmsRaw_TriggerDisplayPreAlarmLOW" : Bool = PLC AlarmsRaw.TriggerDisplayPreAlarmLOW, 100 ms
   "AlarmsRaw_TriggerDisplayAlarmLOW" : Bool = PLC AlarmsRaw.TriggerDisplayAlarmLOW, 100 ms
   "Operation_Operation_ON" : Bool = PLC Operation.Operation_ON, 1 s